'~S001R05CN.Ix.MigWldNoWld - Robot In No Weld MB1[32].3'; 1028 '~Spare MB1[32].4'; 1029 '~S001R05CN.I.WldCtrlCommOk2 - Robot Weld Controller 2 Comm Not OK MB1[32].5'; 1030 '~Spare MB1[32].6'; 1031 '~Spare MB1[32].7'; 1032 '~S001R05CN.I.StudWld2Rdy - Robot Stud Weld Controller 2 Not Ready MB1[32].8'; 1033 '~S001R05CN.I.Rvt2RdyToOperate - Robot Rivet Controller 2 Not Ready MB1[32].9'; 1034 '~S001R05CN.Ix.LaserWldOn - Robot Laser In No Cut MB1[32].10'; 1035 '~S001R05CN.Ix.GlassNotPres - Robot Laser Glass Not Present MB1[32].11'; 1036 '~S001R05CN.Ix.LaserHeadRdy - Robot Laser Head Not Ready MB1[32].12'; 1037 '~S001R05CN.Ix.ChillerOn - Robot Laser Chiller Not On MB1[32].13'; 1038 '~S001R05CN.Ix.GasOn - Robot Gas Not On MB1[32].14'; 1039 '~S001R05 Power Meter Not Ready MB1[32].15'; 1040 '~S001R05 No Wire Present Replace Barrel MB1[32].16'; 1041 '~S001R05 Wire Feeder Fault Timer MB1[32].17'; 1042 '~S001R05CN.Ix.NRFlt - Robot Nut Runner Not Ready MB1[32].18'; 1043 '~Spare MB1[32].19'; 1044 '~S001R05CN.M.WrongRivetAtNose - Remove Wrong Rivet At Nose MB1[32].20'; 1045 '~S001R05CN.M.DisableRbtDrvs - In Rivet Zone But Riveter Not In Auto MB1[32].21'; 1046 '~S001R05CN.I.Rvt1SystemInAuto - Rivet Controller 1 Not In Auto MB1[32].22'; 1047 '~S001R05CN.I.Rvt2SystemInAuto - Rivet Controller 2 Not In Auto MB1[32].23'; 1048 '~S001R05CN.M.RvtC1ReelCtr.DN - Reel Change Required MB1[32].24'; 1049 '~S001R05CN.M.RvtC2ReelCtr.DN - Reel Change Required MB1[32].25'; 1050 '~S001R05CN.M.AbortSkipRemain - SkipRemaining Aborted, Reset At Rbt Controller Is Required MB1[32].26'; 1051 '~Spare MB1[32].27'; 1052 '~Spare MB1[32].28'; 1053 '~Spare MB1[32].29'; 1054 '~Spare MB1[32].30'; 1055 '~Spare MB1[32].31'; 1056 '~Spare MB1[33].0'; 1057 '~Spare MB1[33].1'; 1058 '~Spare MB1[33].2'; 1059 '~Spare MB1[33].3'; 1060 '~Spare MB1[33].4'; 1061 '~Spare MB1[33].5'; 1062 '~Spare MB1[33].6'; 1063 '~Spare MB1[33].7'; 1064 '~Spare MB1[33].8'; 1065 '~Spare MB1[33].9'; 1066 '~Spare MB1[33].10'; 1067 '~Spare MB1[33].11'; 1068 '~Spare MB1[33].12'; 1069 '~Spare MB1[33].13'; 1070 '~Spare MB1[33].14'; 1071 '~Spare MB1[33].15'; 1072 '~Spare MB1[33].16'; 1073 '~Spare MB1[33].17'; 1074 '~Spare MB1[33].18'; 1075 '~Spare MB1[33].19'; 1076 '~Spare MB1[33].20'; 1077 '~Spare MB1[33].21'; 1078 '~Spare MB1[33].22'; 1079 '~Spare MB1[33].23'; 1080 '~Spare MB1[33].24'; 1081 '~Spare MB1[33].25'; 1082 '~Spare MB1[33].26'; 1083 '~Spare MB1[33].27'; 1084 '~Spare MB1[33].28'; 1085 '~Spare MB1[33].29'; 1086 '~Spare MB1[33].30'; 1087 '~Spare MB1[33].31'; 1088 '~Spare MB1[34].0'; 1089 '~Spare MB1[34].1'; 1090 '~Spare MB1[34].2'; 1091 '~Spare MB1[34].3'; 1092 '~Spare MB1[34].4'; 1093 '~Spare MB1[34].5'; 1094 '~Spare MB1[34].6'; 1095 '~Spare MB1[34].7'; 1096 '~Spare MB1[34].8'; 1097 '~Spare MB1[34].9'; 1098 '~Spare MB1[34].10'; 1099 '~Spare MB1[34].11'; 1100 '~Spare MB1[34].12'; 1101 '~Spare MB1[34].13'; 1102 '~Spare MB1[34].14'; 1103 '~Spare MB1[34].15'; 1104 '~Spare MB1[34].16'; 1105 '~Spare MB1[34].17'; 1106 '~Spare MB1[34].18'; 1107 '~Spare MB1[34].19'; 1108 '~Spare MB1[34].20'; 1109 '~Spare MB1[34].21'; 1110 '~Spare MB1[34].22'; 1111 '~Spare MB1[34].23'; 1112 '~Spare MB1[34].24'; 1113 '~Spare MB1[34].25'; 1114 '~Spare MB1[34].26'; 1115 '~Spare MB1[34].27'; 1116 '~Spare MB1[34].28'; 1117 '~Spare MB1[34].29'; 1118 '~Spare MB1[34].30'; 1119 '~Spare MB1[34].31'; 1120 '~Spare MB1[35].0'; 1121 '~Spare MB1[35].1'; 1122 '~Spare MB1[35].2'; 1123 '~Spare MB1[35].3'; 1124 '~Spare MB1[35].4'; 1125 '~Spare MB1[35].5'; 1126 '~Spare MB1[35].6'; 1127 '~Spare MB1[35].7'; 1128 '~Spare MB1[35].8'; 1129 '~Spare MB1[35].9'; 1130 '~Spare MB1[35].10'; 1131 '~Spare MB1[35].11'; 1132 '~Spare MB1[35].12'; 1133 '~Spare MB1[35].13'; 1134 '~Spare MB1[35].14'; 1135 '~Spare MB1[35].15'; 1136 '~Spare MB1[35].16'; 1137 '~Spare MB1[35].17'; 1138 '~Spare MB1[35].18'; 1139 '~Spare MB1[35].19'; 1140 '~Spare MB1[35].20'; 1141 '~Spare MB1[35].21'; 1142 '~Spare MB1[35].22'; 1143 '~Spare MB1[35].23'; 1144 '~Spare MB1[35].24'; 1145 '~Spare MB1[35].25'; 1146 '~Spare MB1[35].26'; 1147 '~Spare MB1[35].27'; 1148 '~Spare MB1[35].28'; 1149 '~Spare MB1[35].29'; 1150 '~Spare MB1[35].30'; 1151 '~Spare MB1[35].31'; 1152 '~S001R06ES1 - S001R06 EtherNet Switch Connection Inhibited MB1[36].0'; 1153 '~Spare MB1[36].1'; 1154 '~Spare MB1[36].2'; 1155 '~Spare MB1[36].3'; 1156 '~Spare MB1[36].4'; 1157 '~Spare MB1[36].5'; 1158 '~Spare MB1[36].6'; 1159 '~Spare MB1[36].7'; 1160 '~Spare MB1[36].8'; 1161 '~Spare MB1[36].9'; 1162 '~Spare MB1[36].10'; 1163 '~Spare MB1[36].11'; 1164 '~Spare MB1[36].12'; 1165 '~Spare MB1[36].13'; 1166 '~Spare MB1[36].14'; 1167 '~Spare MB1[36].15'; 1168 '~Spare MB1[36].16'; 1169 '~S001R06Sfty - Robot E-Stop Depressed MB1[36].17'; 1170 '~S001R06Sfty - Robot Safety Interface Not Enabled MB1[36].18'; 1171 '~S001R06Sfty - Robot DCS Has Been Edited MB1[36].19'; 1172 '~S001R06CN - Robot Controller Connection Inhibited MB1[36].20'; 1173 '~S001R06E#B# - Robot End Effector Module Connection Inhibited MB1[36].21'; 1174 '~S001R06E#B# - Robot End Effector Module Connection Inhibited MB1[36].22'; 1175 '~S001R06E#B# - Robot End Effector Module Connection Inhibited MB1[36].23'; 1176 '~S001R06E#B# - Robot End Effector Module Connection Inhibited MB1[36].24'; 1177 '~S001R06E#B# - Robot End Effector Module Connection Inhibited MB1[36].25'; 1178 '~S001R06E#B# - Robot End Effector Module Connection Inhibited MB1[36].26'; 1179 '~S001R06E#B# - Robot End Effector Module Connection Inhibited MB1[36].27'; 1180 '~S001R06E#B# - Robot End Effector Module Connection Inhibited MB1[36].28'; 1181 '~S001R06E#B# - Robot End Effector Module Connection Inhibited MB1[36].29'; 1182 '~Spare MB1[36].30'; 1183 '~Spare MB1[36].31'; 1184 '~Spare MB1[37].0'; 1185 '~S001R06F#B# - Robot Process I/O Connection Inhibited MB1[37].1'; 1186 '~S001R06F#B# - Robot Process I/O Connection Inhibited MB1[37].2'; 1187 '~S001R06F#B# - Robot Process I/O Connection Inhibited MB1[37].3'; 1188 '~S001R06F#B# - Robot Process I/O Connection Inhibited MB1[37].4'; 1189 '~Spare MB1[37].5'; 1190 '~Spare MB1[37].6'; 1191 '~Spare MB1[37].7'; 1192 '~Spare MB1[37].8'; 1193 '~Spare MB1[37].9'; 1194 '~S001R06CN.I.Safety - Chain Fault MB1[37].10'; 1195 '~S001R06CN.I.AirOn - Robot Air Not On MB1[37].11'; 1196 '~S001R06CN.I.RbtAuto - Robot Not in Auto MB1[37].12'; 1197 '~S001R06CN.M.InTeach - Robot In Teach MB1[37].13'; 1198 '~S001R06CN.I.AtMaintPos - Robot At Maintenace MB1[37].14'; 1199 '~S001R06CN.I.RunEnblInterruptAck - Robot In Hold MB1[37].15'; 1200 '~S001R06CN.M.MaintPosSeld - Robot Maintenance Selected MB1[37].16'; 1201 '~Spare MB1[37].17'; 1202 '~Spare MB1[37].18'; 1203 '~Spare MB1[37].19'; 1204 '~S001R06CN.I.ExtAppCommFlt - Robot Application Communication Fault MB1[37].20'; 1205 '~S001R06CN.M.AbortPickupSeld - Robot Abort Pickup Selected MB1[37].21'; 1206 '~S001R06CN.M.RetFmPounceSeld - Robot Return From Pounce Selected MB1[37].22'; 1207 '~S001R06CN.I.StudWld1 Comm Not OK MB1[37].23'; 1208 '~S001R06CN.I.StudWld2 Comm Not OK MB1[37].24'; 1209 '~S001R06CN.I.WldMode - Robot In No Weld MB1[37].25'; 1210 '~S001R06CN.I.PulledTipBypSS - Robot Pulled Tip Bypass Selected MB1[37].26'; 1211 '~S001R06CN.I.FlowNoFlowSS - Robot In No Flow MB1[37].27'; 1212 '~S001R06CN.I.RvtNoRvtSS - Robot In No Rivet MB1[37].28'; 1213 '~S001R06CN.I.WldCtrlCommOk1 - Robot Weld Controller 1 Comm Not OK MB1[37].29'; 1214 '~S001R06CN.I.WldModeStud - Robot In No Weld Stud MB1[37].30'; 1215 '~S001R06CN.Ix.MigWldNoWld - Robot In No Weld Mig MB1[37].31'; 1216 '~S001R06CN.I.StudWld1Rdy - Robot Stud Weld Controller 1 Not Ready MB1[38].0'; 1217 '~S001R06CN.I.Rvt1RdyToOperate - Robot Rivet Controller 1 Not Ready MB1[38].1'; 1218 '~S001R06CN.Ix.MigRdy - Robot Mig Weld Controller Not Ready MB1[38].2'; 1219 '~S001R06CN.Ix.MigWldNoWld - Robot In No Weld MB1[38].3'; 1220 '~Spare MB1[38].4'; 1221 '~S001R06CN.I.WldCtrlCommOk2 - Robot Weld Controller 2 Comm Not OK MB1[38].5'; 1222 '~Spare MB1[38].6'; 1223 '~Spare MB1[38].7'; 1224 '~S001R06CN.I.StudWld2Rdy - Robot Stud Weld Controller 2 Not Ready MB1[38].8'; 1225 '~S001R06CN.I.Rvt2RdyToOperate - Robot Rivet Controller 2 Not Ready MB1[38].9'; 1226 '~S001R06CN.Ix.LaserWldOn - Robot Laser In No Cut MB1[38].10'; 1227 '~S001R06CN.Ix.GlassNotPres - Robot Laser Glass Not Present MB1[38].11'; 1228 '~S001R06CN.Ix.LaserHeadRdy - Robot Laser Head Not Ready MB1[38].12'; 1229 '~S001R06CN.Ix.ChillerOn - Robot Laser Chiller Not On MB1[38].13'; 1230 '~S001R06CN.Ix.GasOn - Robot Gas Not On MB1[38].14'; 1231 '~S001R06 Power Meter Not Ready MB1[38].15'; 1232 '~S001R06 No Wire Present Replace Barrel MB1[38].16'; 1233 '~S001R06 Wire Feeder Fault Timer MB1[38].17'; 1234 '~S001R06CN.Ix.NRFlt - Robot Nut Runner Not Ready MB1[38].18'; 1235 '~Spare MB1[38].19'; 1236 '~S001R06CN.M.WrongRivetAtNose - Remove Wrong Rivet At Nose MB1[38].20'; 1237 '~S001R06CN.M.DisableRbtDrvs - In Rivet Zone But Riveter Not In Auto MB1[38].21'; 1238 '~S001R06CN.I.Rvt1SystemInAuto - Rivet Controller 1 Not In Auto MB1[38].22'; 1239 '~S001R06CN.I.Rvt2SystemInAuto - Rivet Controller 2 Not In Auto MB1[38].23'; 1240 '~S001R06CN.M.RvtC1ReelCtr.DN - Reel Change Required MB1[38].24'; 1241 '~S001R06CN.M.RvtC2ReelCtr.DN - Reel Change Required MB1[38].25'; 1242 '~S001R06CN.M.AbortSkipRemain - SkipRemaining Aborted, Reset At Rbt Controller Is Required MB1[38].26'; 1243 '~Spare MB1[38].27'; 1244 '~Spare MB1[38].28'; 1245 '~Spare MB1[38].29'; 1246 '~Spare MB1[38].30'; 1247 '~Spare MB1[38].31'; 1248 '~Spare MB1[39].0'; 1249 '~Spare MB1[39].1'; 1250 '~Spare MB1[39].2'; 1251 '~Spare MB1[39].3'; 1252 '~Spare MB1[39].4'; 1253 '~Spare MB1[39].5'; 1254 '~Spare MB1[39].6'; 1255 '~Spare MB1[39].7'; 1256 '~Spare MB1[39].8'; 1257 '~Spare MB1[39].9'; 1258 '~Spare MB1[39].10'; 1259 '~Spare MB1[39].11'; 1260 '~Spare MB1[39].12'; 1261 '~Spare MB1[39].13'; 1262 '~Spare MB1[39].14'; 1263 '~Spare MB1[39].15'; 1264 '~Spare MB1[39].16'; 1265 '~Spare MB1[39].17'; 1266 '~Spare MB1[39].18'; 1267 '~Spare MB1[39].19'; 1268 '~Spare MB1[39].20'; 1269 '~Spare MB1[39].21'; 1270 '~Spare MB1[39].22'; 1271 '~Spare MB1[39].23'; 1272 '~Spare MB1[39].24'; 1273 '~Spare MB1[39].25'; 1274 '~Spare MB1[39].26'; 1275 '~Spare MB1[39].27'; 1276 '~Spare MB1[39].28'; 1277 '~Spare MB1[39].29'; 1278 '~Spare MB1[39].30'; 1279 '~Spare MB1[39].31'; 1280 '~Spare MB1[40].0'; 1281 '~Spare MB1[40].1'; 1282 '~Spare MB1[40].2'; 1283 '~Spare MB1[40].3'; 1284 '~Spare MB1[40].4'; 1285 '~Spare MB1[40].5'; 1286 '~Spare MB1[40].6'; 1287 '~Spare MB1[40].7'; 1288 '~Spare MB1[40].8'; 1289 '~Spare MB1[40].9'; 1290 '~Spare MB1[40].10'; 1291 '~Spare MB1[40].11'; 1292 '~Spare MB1[40].12'; 1293 '~Spare MB1[40].13'; 1294 '~Spare MB1[40].14'; 1295 '~Spare MB1[40].15'; 1296 '~Spare MB1[40].16'; 1297 '~Spare MB1[40].17'; 1298 '~Spare MB1[40].18'; 1299 '~Spare MB1[40].19'; 1300 '~Spare MB1[40].20'; 1301 '~Spare MB1[40].21'; 1302 '~Spare MB1[40].22'; 1303 '~Spare MB1[40].23'; 1304 '~Spare MB1[40].24'; 1305 '~Spare MB1[40].25'; 1306 '~Spare MB1[40].26'; 1307 '~Spare MB1[40].27'; 1308 '~Spare MB1[40].28'; 1309 '~Spare MB1[40].29'; 1310 '~Spare MB1[40].30'; 1311 '~Spare MB1[40].31'; 1312 '~Spare MB1[41].0'; 1313 '~Spare MB1[41].1'; 1314 '~Spare MB1[41].2'; 1315 '~Spare MB1[41].3'; 1316 '~Spare MB1[41].4'; 1317 '~Spare MB1[41].5'; 1318 '~Spare MB1[41].6'; 1319 '~Spare MB1[41].7'; 1320 '~Spare MB1[41].8'; 1321 '~Spare MB1[41].9'; 1322 '~Spare MB1[41].10'; 1323 '~Spare MB1[41].11'; 1324 '~Spare MB1[41].12'; 1325 '~Spare MB1[41].13'; 1326 '~Spare MB1[41].14'; 1327 '~Spare MB1[41].15'; 1328 '~Spare MB1[41].16'; 1329 '~Spare MB1[41].17'; 1330 '~Spare MB1[41].18'; 1331 '~Spare MB1[41].19'; 1332 '~Spare MB1[41].20'; 1333 '~Spare MB1[41].21'; 1334 '~Spare MB1[41].22'; 1335 '~Spare MB1[41].23'; 1336 '~Spare MB1[41].24'; 1337 '~Spare MB1[41].25'; 1338 '~Spare MB1[41].26'; 1339 '~Spare MB1[41].27'; 1340 '~Spare MB1[41].28'; 1341 '~Spare MB1[41].29'; 1342 '~Spare MB1[41].30'; 1343 '~Spare MB1[41].31'; 1344 '~S001R07ES1 - S001R07 EtherNet Switch Connection Inhibited MB1[42].0'; 1345 '~Spare MB1[42].1'; 1346 '~Spare MB1[42].2'; 1347 '~Spare MB1[42].3'; 1348 '~Spare MB1[42].4'; 1349 '~Spare MB1[42].5'; 1350 '~Spare MB1[42].6'; 1351 '~Spare MB1[42].7'; 1352 '~Spare MB1[42].8'; 1353 '~Spare MB1[42].9'; 1354 '~Spare MB1[42].10'; 1355 '~Spare MB1[42].11'; 1356 '~Spare MB1[42].12'; 1357 '~Spare MB1[42].13'; 1358 '~Spare MB1[42].14'; 1359 '~Spare MB1[42].15'; 1360 '~Spare MB1[42].16'; 1361 '~S001R07Sfty - Robot E-Stop Depressed MB1[42].17'; 1362 '~S001R07Sfty - Robot Safety Interface Not Enabled MB1[42].18'; 1363 '~S001R07Sfty - Robot DCS Has Been Edited MB1[42].19'; 1364 '~S001R07CN - Robot Controller Connection Inhibited MB1[42].20'; 1365 '~S001R07E#B# - Robot End Effector Module Connection Inhibited MB1[42].21'; 1366 '~S001R07E#B# - Robot End Effector Module Connection Inhibited MB1[42].22'; 1367 '~S001R07E#B# - Robot End Effector Module Connection Inhibited MB1[42].23'; 1368 '~S001R07E#B# - Robot End Effector Module Connection Inhibited MB1[42].24'; 1369 '~S001R07E#B# - Robot End Effector Module Connection Inhibited MB1[42].25'; 1370 '~S001R07E#B# - Robot End Effector Module Connection Inhibited MB1[42].26'; 1371 '~S001R07E#B# - Robot End Effector Module Connection Inhibited MB1[42].27'; 1372 '~S001R07E#B# - Robot End Effector Module Connection Inhibited MB1[42].28'; 1373 '~S001R07E#B# - Robot End Effector Module Connection Inhibited MB1[42].29'; 1374 '~Spare MB1[42].30'; 1375 '~Spare MB1[42].31'; 1376 '~Spare MB1[43].0'; 1377 '~S001R07F#B# - Robot Process I/O Connection Inhibited MB1[43].1'; 1378 '~S001R07F#B# - Robot Process I/O Connection Inhibited MB1[43].2'; 1379 '~S001R07F#B# - Robot Process I/O Connection Inhibited MB1[43].3'; 1380 '~S001R07F#B# - Robot Process I/O Connection Inhibited MB1[43].4'; 1381 '~Spare MB1[43].5'; 1382 '~Spare MB1[43].6'; 1383 '~Spare MB1[43].7'; 1384 '~Spare MB1[43].8'; 1385 '~Spare MB1[43].9'; 1386 '~S001R07CN.I.Safety - Chain Fault MB1[43].10'; 1387 '~S001R07CN.I.AirOn - Robot Air Not On MB1[43].11'; 1388 '~S001R07CN.I.RbtAuto - Robot Not in Auto MB1[43].12'; 1389 '~S001R07CN.M.InTeach - Robot In Teach MB1[43].13'; 1390 '~S001R07CN.I.AtMaintPos - Robot At Maintenace MB1[43].14'; 1391 '~S001R07CN.I.RunEnblInterruptAck - Robot In Hold MB1[43].15'; 1392 '~S001R07CN.M.MaintPosSeld - Robot Maintenance Selected MB1[43].16'; 1393 '~Spare MB1[43].17'; 1394 '~Spare MB1[43].18'; 1395 '~Spare MB1[43].19'; 1396 '~S001R07CN.I.ExtAppCommFlt - Robot Application Communication Fault MB1[43].20'; 1397 '~S001R07CN.M.AbortPickupSeld - Robot Abort Pickup Selected MB1[43].21'; 1398 '~S001R07CN.M.RetFmPounceSeld - Robot Return From Pounce Selected MB1[43].22'; 1399 '~S001R07CN.I.StudWld1 Comm Not OK MB1[43].23'; 1400 '~S001R07CN.I.StudWld2 Comm Not OK MB1[43].24'; 1401 '~S001R07CN.I.WldMode - Robot In No Weld MB1[43].25'; 1402 '~S001R07CN.I.PulledTipBypSS - Robot Pulled Tip Bypass Selected MB1[43].26'; 1403 '~S001R07CN.I.FlowNoFlowSS - Robot In No Flow MB1[43].27'; 1404 '~S001R07CN.I.RvtNoRvtSS - Robot In No Rivet MB1[43].28'; 1405 '~S001R07CN.I.WldCtrlCommOk1 - Robot Weld Controller 1 Comm Not OK MB1[43].29'; 1406 '~S001R07CN.I.WldModeStud - Robot In No Weld Stud MB1[43].30'; 1407 '~S001R07CN.Ix.MigWldNoWld - Robot In No Weld Mig MB1[43].31'; 1408 '~S001R07CN.I.StudWld1Rdy - Robot Stud Weld Controller 1 Not Ready MB1[44].0'; 1409 '~S001R07CN.I.Rvt1RdyToOperate - Robot Rivet Controller 1 Not Ready MB1[44].1'; 1410 '~S001R07CN.Ix.MigRdy - Robot Mig Weld Controller Not Ready MB1[44].2'; 1411 '~S001R07CN.Ix.MigWldNoWld - Robot In No Weld MB1[44].3'; 1412 '~Spare MB1[44].4'; 1413 '~S001R07CN.I.WldCtrlCommOk2 - Robot Weld Controller 2 Comm Not OK MB1[44].5'; 1414 '~Spare MB1[44].6'; 1415 '~Spare MB1[44].7'; 1416 '~S001R07CN.I.StudWld2Rdy - Robot Stud Weld Controller 2 Not Ready MB1[44].8'; 1417 '~S001R07CN.I.Rvt2RdyToOperate - Robot Rivet Controller 2 Not Ready MB1[44].9'; 1418 '~S001R07CN.Ix.LaserWldOn - Robot Laser In No Cut MB1[44].10'; 1419 '~S001R07CN.Ix.GlassNotPres - Robot Laser Glass Not Present MB1[44].11'; 1420 '~S001R07CN.Ix.LaserHeadRdy - Robot Laser Head Not Ready MB1[44].12'; 1421 '~S001R07CN.Ix.ChillerOn - Robot Laser Chiller Not On MB1[44].13'; 1422 '~S001R07CN.Ix.GasOn - Robot Gas Not On MB1[44].14'; 1423 '~S001R07 Power Meter Not Ready MB1[44].15'; 1424 '~S001R07 No Wire Present Replace Barrel MB1[44].16'; 1425 '~S001R07 Wire Feeder Fault Timer MB1[44].17'; 1426 '~S001R07CN.Ix.NRFlt - Robot Nut Runner Not Ready MB1[44].18'; 1427 '~Spare MB1[44].19'; 1428 '~S001R07CN.M.WrongRivetAtNose - Remove Wrong Rivet At Nose MB1[44].20'; 1429 '~S001R07CN.M.DisableRbtDrvs - In Rivet Zone But Riveter Not In Auto MB1[44].21'; 1430 '~S001R07CN.I.Rvt1SystemInAuto - Rivet Controller 1 Not In Auto MB1[44].22'; 1431 '~S001R07CN.I.Rvt2SystemInAuto - Rivet Controller 2 Not In Auto MB1[44].23'; 1432 '~S001R07CN.M.RvtC1ReelCtr.DN - Reel Change Required MB1[44].24'; 1433 '~S001R07CN.M.RvtC2ReelCtr.DN - Reel Change Required MB1[44].25'; 1434 '~S001R07CN.M.AbortSkipRemain - SkipRemaining Aborted, Reset At Rbt Controller Is Required MB1[44].26'; 1435 '~Spare MB1[44].27'; 1436 '~Spare MB1[44].28'; 1437 '~Spare MB1[44].29'; 1438 '~Spare MB1[44].30'; 1439 '~Spare MB1[44].31'; 1440 '~Spare MB1[45].0'; 1441 '~Spare MB1[45].1'; 1442 '~Spare MB1[45].2'; 1443 '~Spare MB1[45].3'; 1444 '~Spare MB1[45].4'; 1445 '~Spare MB1[45].5'; 1446 '~Spare MB1[45].6'; 1447 '~Spare MB1[45].7'; 1448 '~Spare MB1[45].8'; 1449 '~Spare MB1[45].9'; 1450 '~Spare MB1[45].10'; 1451 '~Spare MB1[45].11'; 1452 '~Spare MB1[45].12'; 1453 '~Spare MB1[45].13'; 1454 '~Spare MB1[45].14'; 1455 '~Spare MB1[45].15'; 1456 '~Spare MB1[45].16'; 1457 '~Spare MB1[45].17'; 1458 '~Spare MB1[45].18'; 1459 '~Spare MB1[45].19'; 1460 '~Spare MB1[45].20'; 1461 '~Spare MB1[45].21'; 1462 '~Spare MB1[45].22'; 1463 '~Spare MB1[45].23'; 1464 '~Spare MB1[45].24'; 1465 '~Spare MB1[45].25'; 1466 '~Spare MB1[45].26'; 1467 '~Spare MB1[45].27'; 1468 '~Spare MB1[45].28'; 1469 '~Spare MB1[45].29'; 1470 '~Spare MB1[45].30'; 1471 '~Spare MB1[45].31'; 1472 '~Spare MB1[46].0'; 1473 '~Spare MB1[46].1'; 1474 '~Spare MB1[46].2'; 1475 '~Spare MB1[46].3'; 1476 '~Spare MB1[46].4'; 1477 '~Spare MB1[46].5'; 1478 '~Spare MB1[46].6'; 1479 '~Spare MB1[46].7'; 1480 '~Spare MB1[46].8'; 1481 '~Spare MB1[46].9'; 1482 '~Spare MB1[46].10'; 1483 '~Spare MB1[46].11'; 1484 '~Spare MB1[46].12'; 1485 '~Spare MB1[46].13'; 1486 '~Spare MB1[46].14'; 1487 '~Spare MB1[46].15'; 1488 '~Spare MB1[46].16'; 1489 '~Spare MB1[46].17'; 1490 '~Spare MB1[46].18'; 1491 '~Spare MB1[46].19'; 1492 '~Spare MB1[46].20'; 1493 '~Spare MB1[46].21'; 1494 '~Spare MB1[46].22'; 1495 '~Spare MB1[46].23'; 1496 '~Spare MB1[46].24'; 1497 '~Spare MB1[46].25'; 1498 '~Spare MB1[46].26'; 1499 '~Spare MB1[46].27'; 1500 '~Spare MB1[46].28'; 1501 '~Spare MB1[46].29'; 1502 '~Spare MB1[46].30'; 1503 '~Spare MB1[46].31'; 1504 '~Spare MB1[47].0'; 1505 '~Spare MB1[47].1'; 1506 '~Spare MB1[47].2'; 1507 '~Spare MB1[47].3'; 1508 '~Spare MB1[47].4'; 1509 '~Spare MB1[47].5'; 1510 '~Spare MB1[47].6'; 1511 '~Spare MB1[47].7'; 1512 '~Spare MB1[47].8'; 1513 '~Spare MB1[47].9'; 1514 '~Spare MB1[47].10'; 1515 '~Spare MB1[47].11'; 1516 '~Spare MB1[47].12'; 1517 '~Spare MB1[47].13'; 1518 '~Spare MB1[47].14'; 1519 '~Spare MB1[47].15'; 1520 '~Spare MB1[47].16'; 1521 '~Spare MB1[47].17'; 1522 '~Spare MB1[47].18'; 1523 '~Spare MB1[47].19'; 1524 '~Spare MB1[47].20'; 1525 '~Spare MB1[47].21'; 1526 '~Spare MB1[47].22'; 1527 '~Spare MB1[47].23'; 1528 '~Spare MB1[47].24'; 1529 '~Spare MB1[47].25'; 1530 '~Spare MB1[47].26'; 1531 '~Spare MB1[47].27'; 1532 '~Spare MB1[47].28'; 1533 '~Spare MB1[47].29'; 1534 '~Spare MB1[47].30'; 1535 '~Spare MB1[47].31'; 1536 '~S001R08ES1 - S001R08 EtherNet Switch Connection Inhibited MB1[48].0'; 1537 '~Spare MB1[48].1'; 1538 '~Spare MB1[48].2'; 1539 '~Spare MB1[48].3'; 1540 '~Spare MB1[48].4'; 1541 '~Spare MB1[48].5'; 1542 '~Spare MB1[48].6'; 1543 '~Spare MB1[48].7'; 1544 '~Spare MB1[48].8'; 1545 '~Spare MB1[48].9'; 1546 '~Spare MB1[48].10'; 1547 '~Spare MB1[48].11'; 1548 '~Spare MB1[48].12'; 1549 '~Spare MB1[48].13'; 1550 '~Spare MB1[48].14'; 1551 '~Spare MB1[48].15'; 1552 '~Spare MB1[48].16'; 1553 '~S001R08Sfty - Robot E-Stop Depressed MB1[48].17'; 1554 '~S001R08Sfty - Robot Safety Interface Not Enabled MB1[48].18'; 1555 '~S001R08Sfty - Robot DCS Has Been Edited MB1[48].19'; 1556 '~S001R08CN - Robot Controller Connection Inhibited MB1[48].20'; 1557 '~S001R08E#B# - Robot End Effector Module Connection Inhibited MB1[48].21'; 1558 '~S001R08E#B# - Robot End Effector Module Connection Inhibited MB1[48].22'; 1559 '~S001R08E#B# - Robot End Effector Module Connection Inhibited MB1[48].23'; 1560 '~S001R08E#B# - Robot End Effector Module Connection Inhibited MB1[48].24'; 1561 '~S001R08E#B# - Robot End Effector Module Connection Inhibited MB1[48].25'; 1562 '~S001R08E#B# - Robot End Effector Module Connection Inhibited MB1[48].26'; 1563 '~S001R08E#B# - Robot End Effector Module Connection Inhibited MB1[48].27'; 1564 '~S001R08E#B# - Robot End Effector Module Connection Inhibited MB1[48].28'; 1565 '~S001R08E#B# - Robot End Effector Module Connection Inhibited MB1[48].29'; 1566 '~Spare MB1[48].30'; 1567 '~Spare MB1[48].31'; 1568 '~Spare MB1[49].0'; 1569 '~S001R08F#B# - Robot Process I/O Connection Inhibited MB1[49].1'; 1570 '~S001R08F#B# - Robot Process I/O Connection Inhibited MB1[49].2'; 1571 '~S001R08F#B# - Robot Process I/O Connection Inhibited MB1[49].3'; 1572 '~S001R08F#B# - Robot Process I/O Connection Inhibited MB1[49].4'; 1573 '~Spare MB1[49].5'; 1574 '~Spare MB1[49].6'; 1575 '~Spare MB1[49].7'; 1576 '~Spare MB1[49].8'; 1577 '~Spare MB1[49].9'; 1578 '~S001R08CN.I.Safety - Chain Fault MB1[49].10'; 1579 '~S001R08CN.I.AirOn - Robot Air Not On MB1[49].11'; 1580 '~S001R08CN.I.RbtAuto - Robot Not in Auto MB1[49].12'; 1581 '~S001R08CN.M.InTeach - Robot In Teach MB1[49].13'; 1582 '~S001R08CN.I.AtMaintPos - Robot At Maintenace MB1[49].14'; 1583 '~S001R08CN.I.RunEnblInterruptAck - Robot In Hold MB1[49].15'; 1584 '~S001R08CN.M.MaintPosSeld - Robot Maintenance Selected MB1[49].16'; 1585 '~Spare MB1[49].17'; 1586 '~Spare MB1[49].18'; 1587 '~Spare MB1[49].19'; 1588 '~S001R08CN.I.ExtAppCommFlt - Robot Application Communication Fault MB1[49].20'; 1589 '~S001R08CN.M.AbortPickupSeld - Robot Abort Pickup Selected MB1[49].21'; 1590 '~S001R08CN.M.RetFmPounceSeld - Robot Return From Pounce Selected MB1[49].22'; 1591 '~S001R08CN.I.StudWld1 Comm Not OK MB1[49].23'; 1592 '~S001R08CN.I.StudWld2 Comm Not OK MB1[49].24'; 1593 '~S001R08CN.I.WldMode - Robot In No Weld MB1[49].25'; 1594 '~S001R08CN.I.PulledTipBypSS - Robot Pulled Tip Bypass Selected MB1[49].26'; 1595 '~S001R08CN.I.FlowNoFlowSS - Robot In No Flow MB1[49].27'; 1596 '~S001R08CN.I.RvtNoRvtSS - Robot In No Rivet MB1[49].28'; 1597 '~S001R08CN.I.WldCtrlCommOk1 - Robot Weld Controller 1 Comm Not OK MB1[49].29'; 1598 '~S001R08CN.I.WldModeStud - Robot In No Weld Stud MB1[49].30'; 1599 '~S001R08CN.Ix.MigWldNoWld - Robot In No Weld Mig MB1[49].31'; 1600 '~S001R08CN.I.StudWld1Rdy - Robot Stud Weld Controller 1 Not Ready MB1[50].0'; 1601 '~S001R08CN.I.Rvt1RdyToOperate - Robot Rivet Controller 1 Not Ready MB1[50].1'; 1602 '~S001R08CN.Ix.MigRdy - Robot Mig Weld Controller Not Ready MB1[50].2'; 1603 '~S001R08CN.Ix.MigWldNoWld - Robot In No Weld MB1[50].3'; 1604 '~Spare MB1[50].4'; 1605 '~S001R08CN.I.WldCtrlCommOk2 - Robot Weld Controller 2 Comm Not OK MB1[50].5'; 1606 '~Spare MB1[50].6'; 1607 '~Spare MB1[50].7'; 1608 '~S001R08CN.I.StudWld2Rdy - Robot Stud Weld Controller 2 Not Ready MB1[50].8'; 1609 '~S001R08CN.I.Rvt2RdyToOperate - Robot Rivet Controller 2 Not Ready MB1[50].9'; 1610 '~S001R08CN.Ix.LaserWldOn - Robot Laser In No Cut MB1[50].10'; 1611 '~S001R08CN.Ix.GlassNotPres - Robot Laser Glass Not Present MB1[50].11'; 1612 '~S001R08CN.Ix.LaserHeadRdy - Robot Laser Head Not Ready MB1[50].12'; 1613 '~S001R08CN.Ix.ChillerOn - Robot Laser Chiller Not On MB1[50].13'; 1614 '~S001R08CN.Ix.GasOn - Robot Gas Not On MB1[50].14'; 1615 '~S001R08 Power Meter Not Ready MB1[50].15'; 1616 '~S001R08 No Wire Present Replace Barrel MB1[50].16'; 1617 '~S001R08 Wire Feeder Fault Timer MB1[50].17'; 1618 '~S001R08CN.Ix.NRFlt - Robot Nut Runner Not Ready MB1[50].18'; 1619 '~Spare MB1[50].19'; 1620 '~S001R08CN.M.WrongRivetAtNose - Remove Wrong Rivet At Nose MB1[50].20'; 1621 '~S001R08CN.M.DisableRbtDrvs - In Rivet Zone But Riveter Not In Auto MB1[50].21'; 1622 '~S001R08CN.I.Rvt1SystemInAuto - Rivet Controller 1 Not In Auto MB1[50].22'; 1623 '~S001R08CN.I.Rvt2SystemInAuto - Rivet Controller 2 Not In Auto MB1[50].23'; 1624 '~S001R08CN.M.RvtC1ReelCtr.DN - Reel Change Required MB1[50].24'; 1625 '~S001R08CN.M.RvtC2ReelCtr.DN - Reel Change Required MB1[50].25'; 1626 '~S001R08CN.M.AbortSkipRemain - SkipRemaining Aborted, Reset At Rbt Controller Is Required MB1[50].26'; 1627 '~Spare MB1[50].27'; 1628 '~Spare MB1[50].28'; 1629 '~Spare MB1[50].29'; 1630 '~Spare MB1[50].30'; 1631 '~Spare MB1[50].31'; 1632 '~Spare MB1[51].0'; 1633 '~Spare MB1[51].1'; 1634 '~Spare MB1[51].2'; 1635 '~Spare MB1[51].3'; 1636 '~Spare MB1[51].4'; 1637 '~Spare MB1[51].5'; 1638 '~Spare MB1[51].6'; 1639 '~Spare MB1[51].7'; 1640 '~Spare MB1[51].8'; 1641 '~Spare MB1[51].9'; 1642 '~Spare MB1[51].10'; 1643 '~Spare MB1[51].11'; 1644 '~Spare MB1[51].12'; 1645 '~Spare MB1[51].13'; 1646 '~Spare MB1[51].14'; 1647 '~Spare MB1[51].15'; 1648 '~Spare MB1[51].16'; 1649 '~Spare MB1[51].17'; 1650 '~Spare MB1[51].18'; 1651 '~Spare MB1[51].19'; 1652 '~Spare MB1[51].20'; 1653 '~Spare MB1[51].21'; 1654 '~Spare MB1[51].22'; 1655 '~Spare MB1[51].23'; 1656 '~Spare MB1[51].24'; 1657 '~Spare MB1[51].25'; 1658 '~Spare MB1[51].26'; 1659 '~Spare MB1[51].27'; 1660 '~Spare MB1[51].28'; 1661 '~Spare MB1[51].29'; 1662 '~Spare MB1[51].30'; 1663 '~Spare MB1[51].31'; 1664 '~Spare MB1[52].0'; 1665 '~Spare MB1[52].1'; 1666 '~Spare MB1[52].2'; 1667 '~Spare MB1[52].3'; 1668 '~Spare MB1[52].4'; 1669 '~Spare MB1[52].5'; 1670 '~Spare MB1[52].6'; 1671 '~Spare MB1[52].7'; 1672 '~Spare MB1[52].8'; 1673 '~Spare MB1[52].9'; 1674 '~Spare MB1[52].10'; 1675 '~Spare MB1[52].11'; 1676 '~Spare MB1[52].12'; 1677 '~Spare MB1[52].13'; 1678 '~Spare MB1[52].14'; 1679 '~Spare MB1[52].15'; 1680 '~Spare MB1[52].16'; 1681 '~Spare MB1[52].17'; 1682 '~Spare MB1[52].18'; 1683 '~Spare MB1[52].19'; 1684 '~Spare MB1[52].20'; 1685 '~Spare MB1[52].21'; 1686 '~Spare MB1[52].22'; 1687 '~Spare MB1[52].23'; 1688 '~Spare MB1[52].24'; 1689 '~Spare MB1[52].25'; 1690 '~Spare MB1[52].26'; 1691 '~Spare MB1[52].27'; 1692 '~Spare MB1[52].28'; 1693 '~Spare MB1[52].29'; 1694 '~Spare MB1[52].30'; 1695 '~Spare MB1[52].31'; 1696 '~Spare MB1[53].0'; 1697 '~Spare MB1[53].1'; 1698 '~Spare MB1[53].2'; 1699 '~Spare MB1[53].3'; 1700 '~Spare MB1[53].4'; 1701 '~Spare MB1[53].5'; 1702 '~Spare MB1[53].6'; 1703 '~Spare MB1[53].7'; 1704 '~Spare MB1[53].8'; 1705 '~Spare MB1[53].9'; 1706 '~Spare MB1[53].10'; 1707 '~Spare MB1[53].11'; 1708 '~Spare MB1[53].12'; 1709 '~Spare MB1[53].13'; 1710 '~Spare MB1[53].14'; 1711 '~Spare MB1[53].15'; 1712 '~Spare MB1[53].16'; 1713 '~Spare MB1[53].17'; 1714 '~Spare MB1[53].18'; 1715 '~Spare MB1[53].19'; 1716 '~Spare MB1[53].20'; 1717 '~Spare MB1[53].21'; 1718 '~Spare MB1[53].22'; 1719 '~Spare MB1[53].23'; 1720 '~Spare MB1[53].24'; 1721 '~Spare MB1[53].25'; 1722 '~Spare MB1[53].26'; 1723 '~Spare MB1[53].27'; 1724 '~Spare MB1[53].28'; 1725 '~Spare MB1[53].29'; 1726 '~Spare MB1[53].30'; 1727 '~Spare MB1[53].31'; 1728 '~Spare MB1[54].0'; 1729 '~Spare MB1[54].1'; 1730 '~Spare MB1[54].2'; 1731 '~Spare MB1[54].3'; 1732 '~Spare MB1[54].4'; 1733 '~Spare MB1[54].5'; 1734 '~Spare MB1[54].6'; 1735 '~Spare MB1[54].7'; 1736 '~Spare MB1[54].8'; 1737 '~Spare MB1[54].9'; 1738 '~Spare MB1[54].10'; 1739 '~Spare MB1[54].11'; 1740 '~Spare MB1[54].12'; 1741 '~Spare MB1[54].13'; 1742 '~Spare MB1[54].14'; 1743 '~Spare MB1[54].15'; 1744 '~Spare MB1[54].16'; 1745 '~Spare MB1[54].17'; 1746 '~Spare MB1[54].18'; 1747 '~Spare MB1[54].19'; 1748 '~Spare MB1[54].20'; 1749 '~Spare MB1[54].21'; 1750 '~Spare MB1[54].22'; 1751 '~Spare MB1[54].23'; 1752 '~Spare MB1[54].24'; 1753 '~Spare MB1[54].25'; 1754 '~Spare MB1[54].26'; 1755 '~Spare MB1[54].27'; 1756 '~Spare MB1[54].28'; 1757 '~Spare MB1[54].29'; 1758 '~Spare MB1[54].30'; 1759 '~Spare MB1[54].31'; 1760 '~Spare MB1[55].0'; 1761 '~Spare MB1[55].1'; 1762 '~Spare MB1[55].2'; 1763 '~Spare MB1[55].3'; 1764 '~Spare MB1[55].4'; 1765 '~Spare MB1[55].5'; 1766 '~Spare MB1[55].6'; 1767 '~Spare MB1[55].7'; 1768 '~Spare MB1[55].8'; 1769 '~Spare MB1[55].9'; 1770 '~Spare MB1[55].10'; 1771 '~Spare MB1[55].11'; 1772 '~Spare MB1[55].12'; 1773 '~Spare MB1[55].13'; 1774 '~Spare MB1[55].14'; 1775 '~Spare MB1[55].15'; 1776 '~Spare MB1[55].16'; 1777 '~Spare MB1[55].17'; 1778 '~Spare MB1[55].18'; 1779 '~Spare MB1[55].19'; 1780 '~Spare MB1[55].20'; 1781 '~Spare MB1[55].21'; 1782 '~Spare MB1[55].22'; 1783 '~Spare MB1[55].23'; 1784 '~Spare MB1[55].24'; 1785 '~Spare MB1[55].25'; 1786 '~Spare MB1[55].26'; 1787 '~Spare MB1[55].27'; 1788 '~Spare MB1[55].28'; 1789 '~Spare MB1[55].29'; 1790 '~Spare MB1[55].30'; 1791 '~Spare MB1[55].31'; 1792 '~Spare MB1[56].0'; 1793 '~Spare MB1[56].1'; 1794 '~S001LS1Sfty - Operator 1 E-Stop Depressed MB1[56].2'; 1795 '~S001LS1Sfty - Operator 2 E-Stop Depressed MB1[56].3'; 1796 '~Spare MB1[56].4'; 1797 '~Spare MB1[56].5'; 1798 '~Spare MB1[56].6'; 1799 '~Spare MB1[56].7'; 1800 '~Spare MB1[56].8'; 1801 '~Spare MB1[56].9'; 1802 '~S001LS1Sfty - Line Access Light Screen Faulted MB1[56].10'; 1803 '~S001LS1Sfty - Operator 1 Light Screen Faulted MB1[56].11'; 1804 '~S001LS1Sfty - Operator 2 Light Screen Faulted MB1[56].12'; 1805 '~S001LS1Sfty - Operator 3 Light Screen Faulted MB1[56].13'; 1806 '~Spare MB1[56].14'; 1807 '~Spare MB1[56].15'; 1808 '~Spare MB1[56].16'; 1809 '~Spare MB1[56].17'; 1810 '~S001LS2Sfty - Operator 1 E-Stop Depressed MB1[56].18'; 1811 '~S001LS2Sfty - Operator 2 E-Stop Depressed MB1[56].19'; 1812 '~Spare MB1[56].20'; 1813 '~Spare MB1[56].21'; 1814 '~Spare MB1[56].22'; 1815 '~Spare MB1[56].23'; 1816 '~Spare MB1[56].24'; 1817 '~Spare MB1[56].25'; 1818 '~S001LS2Sfty - Line Access Light Screen Faulted MB1[56].26'; 1819 '~S001LS2Sfty - Operator 1 Light Screen Faulted MB1[56].27'; 1820 '~S001LS2Sfty - Operator 2 Light Screen Faulted MB1[56].28'; 1821 '~S001LS2Sfty - Operator 3 Light Screen Faulted MB1[56].29'; 1822 '~Spare MB1[56].30'; 1823 '~Spare MB1[56].31'; 1824 '~Spare MB1[57].0'; 1825 '~Spare MB1[57].1'; 1826 '~Spare MB1[57].2'; 1827 '~Spare MB1[57].3'; 1828 '~Spare MB1[57].4'; 1829 '~Spare MB1[57].5'; 1830 '~Spare MB1[57].6'; 1831 '~Spare MB1[57].7'; 1832 '~Spare MB1[57].8'; 1833 '~Spare MB1[57].9'; 1834 '~Spare MB1[57].10'; 1835 '~Spare MB1[57].11'; 1836 '~Spare MB1[57].12'; 1837 '~Spare MB1[57].13'; 1838 '~Spare MB1[57].14'; 1839 '~Spare MB1[57].15'; 1840 '~Spare MB1[57].16'; 1841 '~Spare MB1[57].17'; 1842 '~Spare MB1[57].18'; 1843 '~Spare MB1[57].19'; 1844 '~Spare MB1[57].20'; 1845 '~Spare MB1[57].21'; 1846 '~Spare MB1[57].22'; 1847 '~Spare MB1[57].23'; 1848 '~Spare MB1[57].24'; 1849 '~Spare MB1[57].25'; 1850 '~Spare MB1[57].26'; 1851 '~Spare MB1[57].27'; 1852 '~Spare MB1[57].28'; 1853 '~Spare MB1[57].29'; 1854 '~Spare MB1[57].30'; 1855 '~Spare MB1[57].31'; 1856 '~Spare MB1[58].0'; 1857 '~Spare MB1[58].1'; 1858 '~Spare MB1[58].2'; 1859 '~Spare MB1[58].3'; 1860 '~Spare MB1[58].4'; 1861 '~Spare MB1[58].5'; 1862 '~Spare MB1[58].6'; 1863 '~Spare MB1[58].7'; 1864 '~Spare MB1[58].8'; 1865 '~Spare MB1[58].9'; 1866 '~Spare MB1[58].10'; 1867 '~Spare MB1[58].11'; 1868 '~Spare MB1[58].12'; 1869 '~Spare MB1[58].13'; 1870 '~Spare MB1[58].14'; 1871 '~Spare MB1[58].15'; 1872 '~Spare MB1[58].16'; 1873 '~Spare MB1[58].17'; 1874 '~Spare MB1[58].18'; 1875 '~Spare MB1[58].19'; 1876 '~Spare MB1[58].20'; 1877 '~Spare MB1[58].21'; 1878 '~Spare MB1[58].22'; 1879 '~Spare MB1[58].23'; 1880 '~Spare MB1[58].24'; 1881 '~Spare MB1[58].25'; 1882 '~Spare MB1[58].26'; 1883 '~Spare MB1[58].27'; 1884 '~Spare MB1[58].28'; 1885 '~Spare MB1[58].29'; 1886 '~Spare MB1[58].30'; 1887 '~Spare MB1[58].31'; 1888 '~Spare MB1[59].0'; 1889 '~Spare MB1[59].1'; 1890 '~Spare MB1[59].2'; 1891 '~Spare MB1[59].3'; 1892 '~Spare MB1[59].4'; 1893 '~Spare MB1[59].5'; 1894 '~Spare MB1[59].6'; 1895 '~Spare MB1[59].7'; 1896 '~Spare MB1[59].8'; 1897 '~Spare MB1[59].9'; 1898 '~Spare MB1[59].10'; 1899 '~Spare MB1[59].11'; 1900 '~Spare MB1[59].12'; 1901 '~Spare MB1[59].13'; 1902 '~Spare MB1[59].14'; 1903 '~Spare MB1[59].15'; 1904 '~Spare MB1[59].16'; 1905 '~Spare MB1[59].17'; 1906 '~Spare MB1[59].18'; 1907 '~Spare MB1[59].19'; 1908 '~Spare MB1[59].20'; 1909 '~Spare MB1[59].21'; 1910 '~Spare MB1[59].22'; 1911 '~Spare MB1[59].23'; 1912 '~Spare MB1[59].24'; 1913 '~Spare MB1[59].25'; 1914 '~Spare MB1[59].26'; 1915 '~Spare MB1[59].27'; 1916 '~Spare MB1[59].28'; 1917 '~Spare MB1[59].29'; 1918 '~Spare MB1[59].30'; 1919 '~Spare MB1[59].31'; 1920 '~Spare MB1[60].0'; 1921 '~Spare MB1[60].1'; 1922 '~Spare MB1[60].2'; 1923 '~Spare MB1[60].3'; 1924 '~Spare MB1[60].4'; 1925 '~Spare MB1[60].5'; 1926 '~Spare MB1[60].6'; 1927 '~Spare MB1[60].7'; 1928 '~Spare MB1[60].8'; 1929 '~Spare MB1[60].9'; 1930 '~Spare MB1[60].10'; 1931 '~Spare MB1[60].11'; 1932 '~Spare MB1[60].12'; 1933 '~Spare MB1[60].13'; 1934 '~Spare MB1[60].14'; 1935 '~Spare MB1[60].15'; 1936 '~Spare MB1[60].16'; 1937 '~Spare MB1[60].17'; 1938 '~Spare MB1[60].18'; 1939 '~Spare MB1[60].19'; 1940 '~Spare MB1[60].20'; 1941 '~Spare MB1[60].21'; 1942 '~Spare MB1[60].22'; 1943 '~Spare MB1[60].23'; 1944 '~Spare MB1[60].24'; 1945 '~Spare MB1[60].25'; 1946 '~Spare MB1[60].26'; 1947 '~Spare MB1[60].27'; 1948 '~Spare MB1[60].28'; 1949 '~Spare MB1[60].29'; 1950 '~Spare MB1[60].30'; 1951 '~Spare MB1[60].31'; 1952 '~Spare MB1[61].0'; 1953 '~Spare MB1[61].1'; 1954 '~Spare MB1[61].2'; 1955 '~Spare MB1[61].3'; 1956 '~Spare MB1[61].4'; 1957 '~Spare MB1[61].5'; 1958 '~Spare MB1[61].6'; 1959 '~Spare MB1[61].7'; 1960 '~Spare MB1[61].8'; 1961 '~Spare MB1[61].9'; 1962 '~Spare MB1[61].10'; 1963 '~Spare MB1[61].11'; 1964 '~Spare MB1[61].12'; 1965 '~Spare MB1[61].13'; 1966 '~Spare MB1[61].14'; 1967 '~Spare MB1[61].15'; 1968 '~Spare MB1[61].16'; 1969 '~Spare MB1[61].17'; 1970 '~Spare MB1[61].18'; 1971 '~Spare MB1[61].19'; 1972 '~Spare MB1[61].20'; 1973 '~Spare MB1[61].21'; 1974 '~Spare MB1[61].22'; 1975 '~Spare MB1[61].23'; 1976 '~Spare MB1[61].24'; 1977 '~Spare MB1[61].25'; 1978 '~Spare MB1[61].26'; 1979 '~Spare MB1[61].27'; 1980 '~Spare MB1[61].28'; 1981 '~Spare MB1[61].29'; 1982 '~Spare MB1[61].30'; 1983 '~Spare MB1[61].31'; 1984 '~Spare MB1[62].0'; 1985 '~Spare MB1[62].1'; 1986 '~Spare MB1[62].2'; 1987 '~Spare MB1[62].3'; 1988 '~Spare MB1[62].4'; 1989 '~Spare MB1[62].5'; 1990 '~Spare MB1[62].6'; 1991 '~Spare MB1[62].7'; 1992 '~Spare MB1[62].8'; 1993 '~Spare MB1[62].9'; 1994 '~Spare MB1[62].10'; 1995 '~Spare MB1[62].11'; 1996 '~Spare MB1[62].12'; 1997 '~Spare MB1[62].13'; 1998 '~Spare MB1[62].14'; 1999 '~Spare MB1[62].15'; 2000 '~Spare MB1[62].16'; 2001 '~Spare MB1[62].17'; 2002 '~Spare MB1[62].18'; 2003 '~Spare MB1[62].19'; 2004 '~Spare MB1[62].20'; 2005 '~Spare MB1[62].21'; 2006 '~Spare MB1[62].22'; 2007 '~Spare MB1[62].23'; 2008 '~Spare MB1[62].24'; 2009 '~Spare MB1[62].25'; 2010 '~Spare MB1[62].26'; 2011 '~Spare MB1[62].27'; 2012 '~Spare MB1[62].28'; 2013 '~Spare MB1[62].29'; 2014 '~Spare MB1[62].30'; 2015 '~Spare MB1[62].31'; 2016 '~Spare MB1[63].0'; 2017 '~Spare MB1[63].1'; 2018 '~Spare MB1[63].2'; 2019 '~Spare MB1[63].3'; 2020 '~Spare MB1[63].4'; 2021 '~Spare MB1[63].5'; 2022 '~Spare MB1[63].6'; 2023 '~Spare MB1[63].7'; 2024 '~Spare MB1[63].8'; 2025 '~Spare MB1[63].9'; 2026 '~Spare MB1[63].10'; 2027 '~Spare MB1[63].11'; 2028 '~Spare MB1[63].12'; 2029 '~Spare MB1[63].13'; 2030 '~Spare MB1[63].14'; 2031 '~Spare MB1[63].15'; 2032 '~Spare MB1[63].16'; 2033 '~Spare MB1[63].17'; 2034 '~Spare MB1[63].18'; 2035 '~Spare MB1[63].19'; 2036 '~Spare MB1[63].20'; 2037 '~Spare MB1[63].21'; 2038 '~Spare MB1[63].22'; 2039 '~Spare MB1[63].23'; 2040 '~Spare MB1[63].24'; 2041 '~Spare MB1[63].25'; 2042 '~Spare MB1[63].26'; 2043 '~Spare MB1[63].27'; 2044 '~Spare MB1[63].28'; 2045 '~Spare MB1[63].29'; 2046 '~Spare MB1[63].30'; 2047 '~Spare MB1[63].31'; 2048 '~Spare MB1[64].0'; 2049 '~Spare MB1[64].1'; 2050 '~Spare MB1[64].2'; 2051 '~Spare MB1[64].3'; 2052 '~Spare MB1[64].4'; 2053 '~Spare MB1[64].5'; 2054 '~Spare MB1[64].6'; 2055 '~Spare MB1[64].7'; 2056 '~Spare MB1[64].8'; 2057 '~Spare MB1[64].9'; 2058 '~Spare MB1[64].10'; 2059 '~Spare MB1[64].11'; 2060 '~Spare MB1[64].12'; 2061 '~Spare MB1[64].13'; 2062 '~Spare MB1[64].14'; 2063 '~Spare MB1[64].15'; 2064 '~Spare MB1[64].16'; 2065 '~Spare MB1[64].17'; 2066 '~Spare MB1[64].18'; 2067 '~Spare MB1[64].19'; 2068 '~Spare MB1[64].20'; 2069 '~Spare MB1[64].21'; 2070 '~Spare MB1[64].22'; 2071 '~Spare MB1[64].23'; 2072 '~Spare MB1[64].24'; 2073 '~Spare MB1[64].25'; 2074 '~Spare MB1[64].26'; 2075 '~Spare MB1[64].27'; 2076 '~Spare MB1[64].28'; 2077 '~Spare MB1[64].29'; 2078 '~Spare MB1[64].30'; 2079 '~Spare MB1[64].31'; 2080 '~Spare MB1[65].0'; 2081 '~Spare MB1[65].1'; 2082 '~Spare MB1[65].2'; 2083 '~Spare MB1[65].3'; 2084 '~Spare MB1[65].4'; 2085 '~Spare MB1[65].5'; 2086 '~Spare MB1[65].6'; 2087 '~Spare MB1[65].7'; 2088 '~Spare MB1[65].8'; 2089 '~Spare MB1[65].9'; 2090 '~Spare MB1[65].10'; 2091 '~Spare MB1[65].11'; 2092 '~Spare MB1[65].12'; 2093 '~Spare MB1[65].13'; 2094 '~Spare MB1[65].14'; 2095 '~Spare MB1[65].15'; 2096 '~Spare MB1[65].16'; 2097 '~Spare MB1[65].17'; 2098 '~Spare MB1[65].18'; 2099 '~Spare MB1[65].19'; 2100 '~Spare MB1[65].20'; 2101 '~Spare MB1[65].21'; 2102 '~Spare MB1[65].22'; 2103 '~Spare MB1[65].23'; 2104 '~Spare MB1[65].24'; 2105 '~Spare MB1[65].25'; 2106 '~Spare MB1[65].26'; 2107 '~Spare MB1[65].27'; 2108 '~Spare MB1[65].28'; 2109 '~Spare MB1[65].29'; 2110 '~Spare MB1[65].30'; 2111 '~Spare MB1[65].31'; 2112 '~Spare MB1[66].0'; 2113 '~Spare MB1[66].1'; 2114 '~Spare MB1[66].2'; 2115 '~Spare MB1[66].3'; 2116 '~Spare MB1[66].4'; 2117 '~Spare MB1[66].5'; 2118 '~Spare MB1[66].6'; 2119 '~Spare MB1[66].7'; 2120 '~Spare MB1[66].8'; 2121 '~Spare MB1[66].9'; 2122 '~Spare MB1[66].10'; 2123 '~Spare MB1[66].11'; 2124 '~Spare MB1[66].12'; 2125 '~Spare MB1[66].13'; 2126 '~Spare MB1[66].14'; 2127 '~Spare MB1[66].15'; 2128 '~Spare MB1[66].16'; 2129 '~Spare MB1[66].17'; 2130 '~Spare MB1[66].18'; 2131 '~Spare MB1[66].19'; 2132 '~Spare MB1[66].20'; 2133 '~Spare MB1[66].21'; 2134 '~Spare MB1[66].22'; 2135 '~Spare MB1[66].23'; 2136 '~Spare MB1[66].24'; 2137 '~Spare MB1[66].25'; 2138 '~Spare MB1[66].26'; 2139 '~Spare MB1[66].27'; 2140 '~Spare MB1[66].28'; 2141 '~Spare MB1[66].29'; 2142 '~Spare MB1[66].30'; 2143 '~Spare MB1[66].31'; 2144 '~Spare MB1[67].0'; 2145 '~Spare MB1[67].1'; 2146 '~Spare MB1[67].2'; 2147 '~Spare MB1[67].3'; 2148 '~Spare MB1[67].4'; 2149 '~Spare MB1[67].5'; 2150 '~Spare MB1[67].6'; 2151 '~Spare MB1[67].7'; 2152 '~Spare MB1[67].8'; 2153 '~Spare MB1[67].9'; 2154 '~Spare MB1[67].10'; 2155 '~Spare MB1[67].11'; 2156 '~Spare MB1[67].12'; 2157 '~Spare MB1[67].13'; 2158 '~Spare MB1[67].14'; 2159 '~Spare MB1[67].15'; 2160 '~Spare MB1[67].16'; 2161 '~Spare MB1[67].17'; 2162 '~Spare MB1[67].18'; 2163 '~Spare MB1[67].19'; 2164 '~Spare MB1[67].20'; 2165 '~Spare MB1[67].21'; 2166 '~Spare MB1[67].22'; 2167 '~Spare MB1[67].23'; 2168 '~Spare MB1[67].24'; 2169 '~Spare MB1[67].25'; 2170 '~Spare MB1[67].26'; 2171 '~Spare MB1[67].27'; 2172 '~Spare MB1[67].28'; 2173 '~Spare MB1[67].29'; 2174 '~Spare MB1[67].30'; 2175 '~Spare MB1[67].31'; 2176 '~S001FX1B# - Module Connection Inhibited MB1[68].0'; 2177 '~S001FX1B# - Module Connection Inhibited MB1[68].1'; 2178 '~S001FX1B# - Module Connection Inhibited MB1[68].2'; 2179 '~S001FX1B# - Module Connection Inhibited MB1[68].3'; 2180 '~S001FX1B# - Module Connection Inhibited MB1[68].4'; 2181 '~S001FX1B# - Module Connection Inhibited MB1[68].5'; 2182 '~S001FX1B# - Module Connection Inhibited MB1[68].6'; 2183 '~S001FX1B# - Module Connection Inhibited MB1[68].7'; 2184 '~Spare MB1[68].8'; 2185 '~Spare MB1[68].9'; 2186 '~Spare MB1[68].10'; 2187 '~Spare MB1[68].11'; 2188 '~Spare MB1[68].12'; 2189 '~Spare MB1[68].13'; 2190 '~Spare MB1[68].14'; 2191 